   (* //Move Z256 ALM
   "DB_M256M_Scada".tAlm.tS.tS0 := "DB_Z256_Scada".tAlm.tS.tS0;
   "DB_Z256_Scada".tAlm.tS.tS0.x0 := "DB_Z256_Scada".tAlm.tS.tS0.x0;
   "DB_Z256_Scada".tAlm.tS.tS0.x1 := "DB_Z256_Scada".tAlm.tS.tS0.x1;
   "DB_Z256_Scada".tAlm.tS.tS0.x2 := "DB_Z256_Scada".tAlm.tS.tS0.x2;
   "DB_Z256_Scada".tAlm.tS.tS0.x3 := "DB_Z256_Scada".tAlm.tS.tS0.x3;
   "DB_Z256_Scada".tAlm.tS.tS0.x4 := "DB_Z256_Scada".tAlm.tS.tS0.x4;
   "DB_Z256_Scada".tAlm.tS.tS0.x5 := "DB_Z256_Scada".tAlm.tS.tS0.x5;
   "DB_Z256_Scada".tAlm.tS.tS0.x6 := "DB_Z256_Scada".tAlm.tS.tS0.x6;
   "DB_Z256_Scada".tAlm.tS.tS0.x7 := "DB_Z256_Scada".tAlm.tS.tS0.x7;
   "DB_Z256_Scada".tAlm.tS.tS0.x8 := "DB_Z256_Scada".tAlm.tS.tS0.x8;

   "DB_Z256_Scada".tAlm.tS.tS0.x9 := "DB_Z256_Scada".tAlm.tS.tS0.x9;
   "DB_Z256_Scada".tAlm.tS.tS0.x10 := "DB_Z256_Scada".tAlm.tS.tS0.x10;
   "DB_Z256_Scada".tAlm.tS.tS0.x11 := "DB_Z256_Scada".tAlm.tS.tS0.x11;
   "DB_Z256_Scada".tAlm.tS.tS0.x12 := "DB_Z256_Scada".tAlm.tS.tS0.x12;
   "DB_Z256_Scada".tAlm.tS.tS0.x13 := "DB_Z256_Scada".tAlm.tS.tS0.x13;
   "DB_Z256_Scada".tAlm.tS.tS0.x14 := "DB_Z256_Scada".tAlm.tS.tS0.x14;
   "DB_Z256_Scada".tAlm.tS.tS0.x15 := "DB_Z256_Scada".tAlm.tS.tS0.x15;
   "DB_Z256_Scada".tAlm.tS.tS0.x16 := "DB_Z256_Scada".tAlm.tS.tS0.x16;
   "DB_Z256_Scada".tAlm.tS.tS0.x17 := "DB_Z256_Scada".tAlm.tS.tS0.x17;

   "DB_Z256_Scada".tAlm.tS.tS0.x18 := "DB_Z256_Scada".tAlm.tS.tS0.x18;
   "DB_Z256_Scada".tAlm.tS.tS0.x19 := "DB_Z256_Scada".tAlm.tS.tS0.x19;
   "DB_Z256_Scada".tAlm.tS.tS0.x20 := "DB_Z256_Scada".tAlm.tS.tS0.x20;
   "DB_Z256_Scada".tAlm.tS.tS0.x21 := "DB_Z256_Scada".tAlm.tS.tS0.x21;
   "DB_Z256_Scada".tAlm.tS.tS0.x22 := "DB_Z256_Scada".tAlm.tS.tS0.x22;
   "DB_Z256_Scada".tAlm.tS.tS0.x23 := "DB_Z256_Scada".tAlm.tS.tS0.x23;
   "DB_Z256_Scada".tAlm.tS.tS0.x24 := "DB_Z256_Scada".tAlm.tS.tS0.x24;
   "DB_Z256_Scada".tAlm.tS.tS0.x25 := "DB_Z256_Scada".tAlm.tS.tS0.x25;
   "DB_Z256_Scada".tAlm.tS.tS0.x26 := "DB_Z256_Scada".tAlm.tS.tS0.x26;
   "DB_Z256_Scada".tAlm.tS.tS0.x27 := "DB_Z256_Scada".tAlm.tS.tS0.x27;
   "DB_Z256_Scada".tAlm.tS.tS0.x28 := "DB_Z256_Scada".tAlm.tS.tS0.x28;
   "DB_Z256_Scada".tAlm.tS.tS0.x29 := "DB_Z256_Scada".tAlm.tS.tS0.x29;
   "DB_Z256_Scada".tAlm.tS.tS0.x30 := "DB_Z256_Scada".tAlm.tS.tS0.x30;
   "DB_Z256_Scada".tAlm.tS.tS0.x31 := "DB_Z256_Scada".tAlm.tS.tS0.x31; *)


    //Move M256M MOVEMENTS HMR
    //H1
   "DB_M256M_Scada".tHMR.tManCmd.xManJogForwardFdbk_H1 := "M256_Manag_IDB".M256M_IDB[0].tHMR.tManCmd.xMan_JogForwardFdbk;
   "DB_M256M_Scada".tHMR.tManCmd.xManJogBackwardFdbk_H1 := "M256_Manag_IDB".M256M_IDB[0].tHMR.tManCmd.xMan_JogBackwardFdbk;
   "DB_M256M_Scada".tHMR.iCodeAlarm_H1 := "M256_Manag_IDB".M256M_IDB[0].tHMR.iCodeAlarm;
   "DB_M256M_Scada".tHMR.dHeadActualPositions_cmm_H1 := "M256_Manag_IDB".M256M_IDB[0].tHMR.dHeadActualPositions_cmm;
   "DB_M256M_Scada".tHMR.dHeadHomePositions_cmm_H1 := "M256_Manag_IDB".M256M_IDB[0].tHMR.dHeadHomePositions_cmm;
   "DB_M256M_Scada".tHMR.dHeadMoveStatus_H1 := "M256_Manag_IDB".M256M_IDB[0].tHMR.rgdHeadMoveStatus;
   //H2 
   "DB_M256M_Scada".tHMR.tManCmd.xManJogBackwardFdbk_H2 := "M256_Manag_IDB".M256M_IDB[1].tHMR.tManCmd.xMan_JogForwardFdbk;
   "DB_M256M_Scada".tHMR.tManCmd.xManJogBackwardFdbk_H2 := "M256_Manag_IDB".M256M_IDB[1].tHMR.tManCmd.xMan_JogBackwardFdbk;
   "DB_M256M_Scada".tHMR.iCodeAlarm_H2 := "M256_Manag_IDB".M256M_IDB[1].tHMR.iCodeAlarm;
   "DB_M256M_Scada".tHMR.dHeadActualPositions_cmm_H2 := "M256_Manag_IDB".M256M_IDB[1].tHMR.dHeadActualPositions_cmm;
   "DB_M256M_Scada".tHMR.dHeadHomePositions_cmm_H2 := "M256_Manag_IDB".M256M_IDB[1].tHMR.dHeadHomePositions_cmm;
   "DB_M256M_Scada".tHMR.dHeadMoveStatus_H2 := "M256_Manag_IDB".M256M_IDB[1].tHMR.rgdHeadMoveStatus;
   //H3 
   "DB_M256M_Scada".tHMR.tManCmd.xManJogForwardFdbk_H3 :="M256_Manag_IDB".M256M_IDB[2].tHMR.tManCmd.xMan_JogForwardFdbk;
   "DB_M256M_Scada".tHMR.tManCmd.xManJogBackwardFdbk_H3 := "M256_Manag_IDB".M256M_IDB[2].tHMR.tManCmd.xMan_JogBackwardFdbk;
   "DB_M256M_Scada".tHMR.iCodeAlarm_H3 := "M256_Manag_IDB".M256M_IDB[2].tHMR.iCodeAlarm;
   "DB_M256M_Scada".tHMR.dHeadActualPositions_cmm_H3 := "M256_Manag_IDB".M256M_IDB[2].tHMR.dHeadActualPositions_cmm;
   "DB_M256M_Scada".tHMR.dHeadHomePositions_cmm_H3 := "M256_Manag_IDB".M256M_IDB[2].tHMR.dHeadHomePositions_cmm;
   "DB_M256M_Scada".tHMR.dHeadMoveStatus_H3 := "M256_Manag_IDB".M256M_IDB[2].tHMR.rgdHeadMoveStatus;
   //H4 
   "DB_M256M_Scada".tHMR.tManCmd.xManJogForwardFdbk_H4:= "M256_Manag_IDB".M256M_IDB[3].tHMR.tManCmd.xMan_JogForwardFdbk;
   "DB_M256M_Scada".tHMR.tManCmd.xManJogBackwardFdbk_H4 := "M256_Manag_IDB".M256M_IDB[3].tHMR.tManCmd.xMan_JogBackwardFdbk;
   "DB_M256M_Scada".tHMR.iCodeAlarm_H4 := "M256_Manag_IDB".M256M_IDB[3].tHMR.iCodeAlarm;
   "DB_M256M_Scada".tHMR.dHeadActualPositions_cmm_H4 := "M256_Manag_IDB".M256M_IDB[3].tHMR.dHeadActualPositions_cmm;
   "DB_M256M_Scada".tHMR.dHeadHomePositions_cmm_H4 := "M256_Manag_IDB".M256M_IDB[3].tHMR.dHeadHomePositions_cmm;
   "DB_M256M_Scada".tHMR.dHeadMoveStatus_H4 := "M256_Manag_IDB".M256M_IDB[3].tHMR.rgdHeadMoveStatus;
   "DB_M256M_Scada".tHMR.iCodeAlarm_H4 := "M256_Manag_IDB".M256M_IDB[3].tHMR.iCodeAlarm;
   //H5
   "DB_M256M_Scada".tHMR.tManCmd.xManJogForwardFdbk_H5 := "M256_Manag_IDB".M256M_IDB[4].tHMR.tManCmd.xMan_JogForwardFdbk;
   "DB_M256M_Scada".tHMR.tManCmd.xManJogBackwardFdbk_H5:= "M256_Manag_IDB".M256M_IDB[4].tHMR.tManCmd.xMan_JogBackwardFdbk;
   "DB_M256M_Scada".tHMR.iCodeAlarm_H5 := "M256_Manag_IDB".M256M_IDB[4].tHMR.iCodeAlarm;
   "DB_M256M_Scada".tHMR.dHeadActualPositions_cmm_H5 := "M256_Manag_IDB".M256M_IDB[4].tHMR.dHeadActualPositions_cmm;
   "DB_M256M_Scada".tHMR.dHeadHomePositions_cmm_H5 := "M256_Manag_IDB".M256M_IDB[4].tHMR.dHeadHomePositions_cmm;
   "DB_M256M_Scada".tHMR.dHeadMoveStatus_H5 := "M256_Manag_IDB".M256M_IDB[4].tHMR.rgdHeadMoveStatus;
   //H6 
   "DB_M256M_Scada".tHMR.tManCmd.xManJogForwardFdbk_H6 := "M256_Manag_IDB".M256M_IDB[5].tHMR.tManCmd.xMan_JogForwardFdbk;
   "DB_M256M_Scada".tHMR.tManCmd.xManJogBackwardFdbk_H6 := "M256_Manag_IDB".M256M_IDB[5].tHMR.tManCmd.xMan_JogBackwardFdbk;
   "DB_M256M_Scada".tHMR.iCodeAlarm_H6 := "M256_Manag_IDB".M256M_IDB[5].tHMR.iCodeAlarm;
   "DB_M256M_Scada".tHMR.dHeadActualPositions_cmm_H6 := "M256_Manag_IDB".M256M_IDB[5].tHMR.dHeadActualPositions_cmm;
   "DB_M256M_Scada".tHMR.dHeadHomePositions_cmm_H6 := "M256_Manag_IDB".M256M_IDB[5].tHMR.dHeadHomePositions_cmm;
   "DB_M256M_Scada".tHMR.dHeadMoveStatus_H6 := "M256_Manag_IDB".M256M_IDB[5].tHMR.rgdHeadMoveStatus;
   //H7 
   "DB_M256M_Scada".tHMR.tManCmd.xManJogForwardFdbk_H7 := "M256_Manag_IDB".M256M_IDB[6].tHMR.tManCmd.xMan_JogForwardFdbk;
   "DB_M256M_Scada".tHMR.tManCmd.xManJogBackwardFdbk_H7 := "M256_Manag_IDB".M256M_IDB[6].tHMR.tManCmd.xMan_JogBackwardFdbk;
   "DB_M256M_Scada".tHMR.iCodeAlarm_H7 := "M256_Manag_IDB".M256M_IDB[6].tHMR.iCodeAlarm;
   "DB_M256M_Scada".tHMR.dHeadActualPositions_cmm_H7 := "M256_Manag_IDB".M256M_IDB[6].tHMR.dHeadActualPositions_cmm;
   "DB_M256M_Scada".tHMR.dHeadHomePositions_cmm_H7 := "M256_Manag_IDB".M256M_IDB[6].tHMR.dHeadHomePositions_cmm;
   "DB_M256M_Scada".tHMR.dHeadMoveStatus_H7 := "M256_Manag_IDB".M256M_IDB[6].tHMR.rgdHeadMoveStatus;
   //H8 
   "DB_M256M_Scada".tHMR.tManCmd.xManJogForwardFdbk_H8 := "M256_Manag_IDB".M256M_IDB[7].tHMR.tManCmd.xMan_JogForwardFdbk;
   "DB_M256M_Scada".tHMR.tManCmd.xManJogBackwardFdbk_H8 := "M256_Manag_IDB".M256M_IDB[7].tHMR.tManCmd.xMan_JogBackwardFdbk;
   "DB_M256M_Scada".tHMR.iCodeAlarm_H8 := "M256_Manag_IDB".M256M_IDB[7].tHMR.iCodeAlarm;
   "DB_M256M_Scada".tHMR.dHeadActualPositions_cmm_H8 := "M256_Manag_IDB".M256M_IDB[7].tHMR.dHeadActualPositions_cmm;
   "DB_M256M_Scada".tHMR.dHeadHomePositions_cmm_H8 := "M256_Manag_IDB".M256M_IDB[7].tHMR.dHeadHomePositions_cmm;
   "DB_M256M_Scada".tHMR.dHeadMoveStatus_H8 := "M256_Manag_IDB".M256M_IDB[7].tHMR.rgdHeadMoveStatus;


       //Move MOVEMENTS HMW

       //H1
       "M256_Manag_IDB".M256M_IDB[0].tHMW.dHeadHomePositions_cmm := "DB_M256M_Scada".tHMW.dHeadHomePositions_cmm_H1;
       "M256_Manag_IDB".M256M_IDB[0].tHMW.xBrakeEngageHeads := "DB_M256M_Scada".tHMW.xBrakeRealeaseHead_H1;
       "M256_Manag_IDB".M256M_IDB[0].tHMW.xBrakeRealeaseHeads := "DB_M256M_Scada".tHMW.xBrakeEngageHeads_H1;
       "M256_Manag_IDB".M256M_IDB[0].tHMW.xUpdateHomeHead := "DB_M256M_Scada".tHMW.xUpdateHomeHead_H1;
       "M256_Manag_IDB".M256M_IDB[0].tHMW.tManCmd.xMan_JogBackward := "DB_M256M_Scada".tHMW.tManCmd.xMan_JogBackward_H1;
       "M256_Manag_IDB".M256M_IDB[0].tHMW.tManCmd.xMan_JogForward := "DB_M256M_Scada".tHMW.tManCmd.xMan_JogForward_H1;
       //H2
       "M256_Manag_IDB".M256M_IDB[1].tHMW.dHeadHomePositions_cmm := "DB_M256M_Scada".tHMW.dHeadHomePositions_cmm_H2;
       "M256_Manag_IDB".M256M_IDB[1].tHMW.xBrakeEngageHeads := "DB_M256M_Scada".tHMW.xBrakeRealeaseHead_H2;
       "M256_Manag_IDB".M256M_IDB[1].tHMW.xBrakeRealeaseHeads := "DB_M256M_Scada".tHMW.xBrakeEngageHeads_H2;
       "M256_Manag_IDB".M256M_IDB[1].tHMW.xUpdateHomeHead := "DB_M256M_Scada".tHMW.xUpdateHomeHead_H2;
       "M256_Manag_IDB".M256M_IDB[1].tHMW.tManCmd.xMan_JogBackward := "DB_M256M_Scada".tHMW.tManCmd.xMan_JogBackward_H2;
       "M256_Manag_IDB".M256M_IDB[1].tHMW.tManCmd.xMan_JogForward := "DB_M256M_Scada".tHMW.tManCmd.xMan_JogForward_H2;
       //H3
       "M256_Manag_IDB".M256M_IDB[2].tHMW.dHeadHomePositions_cmm := "DB_M256M_Scada".tHMW.dHeadHomePositions_cmm_H3;
       "M256_Manag_IDB".M256M_IDB[2].tHMW.xBrakeEngageHeads := "DB_M256M_Scada".tHMW.xBrakeRealeaseHead_H3;
       "M256_Manag_IDB".M256M_IDB[2].tHMW.xBrakeRealeaseHeads := "DB_M256M_Scada".tHMW.xBrakeEngageHeads_H3;
       "M256_Manag_IDB".M256M_IDB[2].tHMW.xUpdateHomeHead := "DB_M256M_Scada".tHMW.xUpdateHomeHead_H3;
       "M256_Manag_IDB".M256M_IDB[2].tHMW.tManCmd.xMan_JogBackward := "DB_M256M_Scada".tHMW.tManCmd.xMan_JogBackward_H3;
       "M256_Manag_IDB".M256M_IDB[2].tHMW.tManCmd.xMan_JogForward := "DB_M256M_Scada".tHMW.tManCmd.xMan_JogForward_H3;
       //H4
       "M256_Manag_IDB".M256M_IDB[3].tHMW.dHeadHomePositions_cmm := "DB_M256M_Scada".tHMW.dHeadHomePositions_cmm_H4;
       "M256_Manag_IDB".M256M_IDB[3].tHMW.xBrakeEngageHeads := "DB_M256M_Scada".tHMW.xBrakeRealeaseHead_H4;
       "M256_Manag_IDB".M256M_IDB[3].tHMW.xBrakeRealeaseHeads := "DB_M256M_Scada".tHMW.xBrakeEngageHeads_H4;
       "M256_Manag_IDB".M256M_IDB[3].tHMW.xUpdateHomeHead := "DB_M256M_Scada".tHMW.xUpdateHomeHead_H4;
       "M256_Manag_IDB".M256M_IDB[3].tHMW.tManCmd.xMan_JogBackward := "DB_M256M_Scada".tHMW.tManCmd.xMan_JogBackward_H4;
       "M256_Manag_IDB".M256M_IDB[3].tHMW.tManCmd.xMan_JogForward := "DB_M256M_Scada".tHMW.tManCmd.xMan_JogForward_H4;
       //H5
       "M256_Manag_IDB".M256M_IDB[4].tHMW.dHeadHomePositions_cmm := "DB_M256M_Scada".tHMW.dHeadHomePositions_cmm_H5;
       "M256_Manag_IDB".M256M_IDB[4].tHMW.xBrakeEngageHeads := "DB_M256M_Scada".tHMW.xBrakeRealeaseHead_H5;
       "M256_Manag_IDB".M256M_IDB[4].tHMW.xBrakeRealeaseHeads := "DB_M256M_Scada".tHMW.xBrakeEngageHeads_H5;
       "M256_Manag_IDB".M256M_IDB[4].tHMW.xUpdateHomeHead := "DB_M256M_Scada".tHMW.xUpdateHomeHead_H5;
       "M256_Manag_IDB".M256M_IDB[4].tHMW.tManCmd.xMan_JogBackward := "DB_M256M_Scada".tHMW.tManCmd.xMan_JogBackward_H5;
       "M256_Manag_IDB".M256M_IDB[4].tHMW.tManCmd.xMan_JogForward := "DB_M256M_Scada".tHMW.tManCmd.xMan_JogForward_H5;
       //H6
       "M256_Manag_IDB".M256M_IDB[5].tHMW.dHeadHomePositions_cmm := "DB_M256M_Scada".tHMW.dHeadHomePositions_cmm_H6;
       "M256_Manag_IDB".M256M_IDB[5].tHMW.xBrakeEngageHeads := "DB_M256M_Scada".tHMW.xBrakeRealeaseHead_H6;
       "M256_Manag_IDB".M256M_IDB[5].tHMW.xBrakeRealeaseHeads := "DB_M256M_Scada".tHMW.xBrakeEngageHeads_H6;
       "M256_Manag_IDB".M256M_IDB[5].tHMW.xUpdateHomeHead := "DB_M256M_Scada".tHMW.xUpdateHomeHead_H6;
       "M256_Manag_IDB".M256M_IDB[5].tHMW.tManCmd.xMan_JogBackward := "DB_M256M_Scada".tHMW.tManCmd.xMan_JogBackward_H6;
       "M256_Manag_IDB".M256M_IDB[5].tHMW.tManCmd.xMan_JogForward := "DB_M256M_Scada".tHMW.tManCmd.xMan_JogForward_H6;
       //H7
       "M256_Manag_IDB".M256M_IDB[6].tHMW.dHeadHomePositions_cmm := "DB_M256M_Scada".tHMW.dHeadHomePositions_cmm_H7;
       "M256_Manag_IDB".M256M_IDB[6].tHMW.xBrakeEngageHeads := "DB_M256M_Scada".tHMW.xBrakeRealeaseHead_H7;
       "M256_Manag_IDB".M256M_IDB[6].tHMW.xBrakeRealeaseHeads := "DB_M256M_Scada".tHMW.xBrakeEngageHeads_H7;
       "M256_Manag_IDB".M256M_IDB[6].tHMW.xUpdateHomeHead := "DB_M256M_Scada".tHMW.xUpdateHomeHead_H7;
       "M256_Manag_IDB".M256M_IDB[6].tHMW.tManCmd.xMan_JogBackward := "DB_M256M_Scada".tHMW.tManCmd.xMan_JogBackward_H7;
       "M256_Manag_IDB".M256M_IDB[6].tHMW.tManCmd.xMan_JogForward := "DB_M256M_Scada".tHMW.tManCmd.xMan_JogForward_H7;

       //H8
       "M256_Manag_IDB".M256M_IDB[7].tHMW.dHeadHomePositions_cmm := "DB_M256M_Scada".tHMW.dHeadHomePositions_cmm_H8;
       "M256_Manag_IDB".M256M_IDB[7].tHMW.xBrakeEngageHeads := "DB_M256M_Scada".tHMW.xBrakeRealeaseHead_H8;
       "M256_Manag_IDB".M256M_IDB[7].tHMW.xBrakeRealeaseHeads := "DB_M256M_Scada".tHMW.xBrakeEngageHeads_H8;
       "M256_Manag_IDB".M256M_IDB[7].tHMW.xUpdateHomeHead := "DB_M256M_Scada".tHMW.xUpdateHomeHead_H8;
       "M256_Manag_IDB".M256M_IDB[7].tHMW.tManCmd.xMan_JogBackward := "DB_M256M_Scada".tHMW.tManCmd.xMan_JogBackward_H8;
       "M256_Manag_IDB".M256M_IDB[7].tHMW.tManCmd.xMan_JogForward := "DB_M256M_Scada".tHMW.tManCmd.xMan_JogForward_H8;

       //Move MOVEMENTS ALM
       //H1
       "DB_M256M_Scada".tAlm.tS.tS0.x0 := "M256_Manag_IDB".M256M_IDB[0].tALM.tS.x0;
       "DB_M256M_Scada".tAlm.tS.tS0.x1 := "M256_Manag_IDB".M256M_IDB[0].tALM.tS.x1;
       "DB_M256M_Scada".tAlm.tS.tS0.x2 := "M256_Manag_IDB".M256M_IDB[0].tALM.tS.x2;
       "DB_M256M_Scada".tAlm.tS.tS0.x3 := "M256_Manag_IDB".M256M_IDB[0].tALM.tS.x3;
       "DB_M256M_Scada".tAlm.tS.tS0.x4 := "M256_Manag_IDB".M256M_IDB[0].tALM.tS.x4;
       "DB_M256M_Scada".tAlm.tS.tS0.x5 := "M256_Manag_IDB".M256M_IDB[0].tALM.tS.x5;
       "DB_M256M_Scada".tAlm.tS.tS0.x6 := "M256_Manag_IDB".M256M_IDB[0].tALM.tS.x6;
       "DB_M256M_Scada".tAlm.tS.tS0.x7 := "M256_Manag_IDB".M256M_IDB[0].tALM.tS.x7;
       "DB_M256M_Scada".tAlm.tS.tS0.x8 := "M256_Manag_IDB".M256M_IDB[0].tALM.tS.x8;
       //H2
       "DB_M256M_Scada".tAlm.tS.tS0.x9 := "M256_Manag_IDB".M256M_IDB[1].tALM.tS.x0;
       "DB_M256M_Scada".tAlm.tS.tS0.x10 := "M256_Manag_IDB".M256M_IDB[1].tALM.tS.x1;
       "DB_M256M_Scada".tAlm.tS.tS0.x11 := "M256_Manag_IDB".M256M_IDB[1].tALM.tS.x2;
       "DB_M256M_Scada".tAlm.tS.tS0.x12 := "M256_Manag_IDB".M256M_IDB[1].tALM.tS.x3;
       "DB_M256M_Scada".tAlm.tS.tS0.x13 := "M256_Manag_IDB".M256M_IDB[1].tALM.tS.x4;
       "DB_M256M_Scada".tAlm.tS.tS0.x14 := "M256_Manag_IDB".M256M_IDB[1].tALM.tS.x5;
       "DB_M256M_Scada".tAlm.tS.tS0.x15 := "M256_Manag_IDB".M256M_IDB[1].tALM.tS.x6;
       "DB_M256M_Scada".tAlm.tS.tS0.x16 := "M256_Manag_IDB".M256M_IDB[1].tALM.tS.x7;
       "DB_M256M_Scada".tAlm.tS.tS0.x17 := "M256_Manag_IDB".M256M_IDB[1].tALM.tS.x8;
       //H3
       "DB_M256M_Scada".tAlm.tS.tS0.x18 := "M256_Manag_IDB".M256M_IDB[2].tALM.tS.x0;
       "DB_M256M_Scada".tAlm.tS.tS0.x19 := "M256_Manag_IDB".M256M_IDB[2].tALM.tS.x1;
       "DB_M256M_Scada".tAlm.tS.tS0.x20 := "M256_Manag_IDB".M256M_IDB[2].tALM.tS.x2;
       "DB_M256M_Scada".tAlm.tS.tS0.x21 := "M256_Manag_IDB".M256M_IDB[2].tALM.tS.x3;
       "DB_M256M_Scada".tAlm.tS.tS0.x22 := "M256_Manag_IDB".M256M_IDB[2].tALM.tS.x4;
       "DB_M256M_Scada".tAlm.tS.tS0.x23 := "M256_Manag_IDB".M256M_IDB[2].tALM.tS.x5;
       "DB_M256M_Scada".tAlm.tS.tS0.x24 := "M256_Manag_IDB".M256M_IDB[2].tALM.tS.x6;
       "DB_M256M_Scada".tAlm.tS.tS0.x25 := "M256_Manag_IDB".M256M_IDB[2].tALM.tS.x7;
       "DB_M256M_Scada".tAlm.tS.tS0.x26 := "M256_Manag_IDB".M256M_IDB[2].tALM.tS.x8;
       //H4
       "DB_M256M_Scada".tAlm.tS.tS1.x0 := "M256_Manag_IDB".M256M_IDB[3].tALM.tS.x0;
       "DB_M256M_Scada".tAlm.tS.tS1.x1 := "M256_Manag_IDB".M256M_IDB[3].tALM.tS.x1;
       "DB_M256M_Scada".tAlm.tS.tS1.x2 := "M256_Manag_IDB".M256M_IDB[3].tALM.tS.x2;
       "DB_M256M_Scada".tAlm.tS.tS1.x3 := "M256_Manag_IDB".M256M_IDB[3].tALM.tS.x3;
       "DB_M256M_Scada".tAlm.tS.tS1.x4 := "M256_Manag_IDB".M256M_IDB[3].tALM.tS.x4;
       "DB_M256M_Scada".tAlm.tS.tS1.x5 := "M256_Manag_IDB".M256M_IDB[3].tALM.tS.x5;
       "DB_M256M_Scada".tAlm.tS.tS1.x6 := "M256_Manag_IDB".M256M_IDB[3].tALM.tS.x6;
       "DB_M256M_Scada".tAlm.tS.tS1.x7 := "M256_Manag_IDB".M256M_IDB[3].tALM.tS.x7;
       "DB_M256M_Scada".tAlm.tS.tS1.x8 := "M256_Manag_IDB".M256M_IDB[3].tALM.tS.x8;
       //H5
       "DB_M256M_Scada".tAlm.tS.tS1.x9 := "M256_Manag_IDB".M256M_IDB[4].tALM.tS.x0;
       "DB_M256M_Scada".tAlm.tS.tS1.x10 := "M256_Manag_IDB".M256M_IDB[4].tALM.tS.x1;
       "DB_M256M_Scada".tAlm.tS.tS1.x11 := "M256_Manag_IDB".M256M_IDB[4].tALM.tS.x2;
       "DB_M256M_Scada".tAlm.tS.tS1.x12 := "M256_Manag_IDB".M256M_IDB[4].tALM.tS.x3;
       "DB_M256M_Scada".tAlm.tS.tS1.x13 := "M256_Manag_IDB".M256M_IDB[4].tALM.tS.x4;
       "DB_M256M_Scada".tAlm.tS.tS1.x14 := "M256_Manag_IDB".M256M_IDB[4].tALM.tS.x5;
       "DB_M256M_Scada".tAlm.tS.tS1.x15 := "M256_Manag_IDB".M256M_IDB[4].tALM.tS.x6;
       "DB_M256M_Scada".tAlm.tS.tS1.x16 := "M256_Manag_IDB".M256M_IDB[4].tALM.tS.x7;
       "DB_M256M_Scada".tAlm.tS.tS1.x17 := "M256_Manag_IDB".M256M_IDB[4].tALM.tS.x8;
       //H6
       "DB_M256M_Scada".tAlm.tS.tS1.x18 := "M256_Manag_IDB".M256M_IDB[5].tALM.tS.x0;
       "DB_M256M_Scada".tAlm.tS.tS1.x19 := "M256_Manag_IDB".M256M_IDB[5].tALM.tS.x1;
       "DB_M256M_Scada".tAlm.tS.tS1.x20 := "M256_Manag_IDB".M256M_IDB[5].tALM.tS.x2;
       "DB_M256M_Scada".tAlm.tS.tS1.x21 := "M256_Manag_IDB".M256M_IDB[5].tALM.tS.x3;
       "DB_M256M_Scada".tAlm.tS.tS1.x22 := "M256_Manag_IDB".M256M_IDB[5].tALM.tS.x4;
       "DB_M256M_Scada".tAlm.tS.tS1.x23 := "M256_Manag_IDB".M256M_IDB[5].tALM.tS.x5;
       "DB_M256M_Scada".tAlm.tS.tS1.x24 := "M256_Manag_IDB".M256M_IDB[5].tALM.tS.x6;
       "DB_M256M_Scada".tAlm.tS.tS1.x25 := "M256_Manag_IDB".M256M_IDB[5].tALM.tS.x7;
       "DB_M256M_Scada".tAlm.tS.tS1.x26 := "M256_Manag_IDB".M256M_IDB[5].tALM.tS.x8;
       //H7
       "DB_M256M_Scada".tAlm.tS.tS2.x0 := "M256_Manag_IDB".M256M_IDB[6].tALM.tS.x0;
       "DB_M256M_Scada".tAlm.tS.tS2.x1 := "M256_Manag_IDB".M256M_IDB[6].tALM.tS.x1;
       "DB_M256M_Scada".tAlm.tS.tS2.x2 := "M256_Manag_IDB".M256M_IDB[6].tALM.tS.x2;
       "DB_M256M_Scada".tAlm.tS.tS2.x3 := "M256_Manag_IDB".M256M_IDB[6].tALM.tS.x3;
       "DB_M256M_Scada".tAlm.tS.tS2.x4 := "M256_Manag_IDB".M256M_IDB[6].tALM.tS.x4;
       "DB_M256M_Scada".tAlm.tS.tS2.x5 := "M256_Manag_IDB".M256M_IDB[6].tALM.tS.x5;
       "DB_M256M_Scada".tAlm.tS.tS2.x6 := "M256_Manag_IDB".M256M_IDB[6].tALM.tS.x6;
       "DB_M256M_Scada".tAlm.tS.tS2.x7 := "M256_Manag_IDB".M256M_IDB[6].tALM.tS.x7;
       "DB_M256M_Scada".tAlm.tS.tS2.x8 := "M256_Manag_IDB".M256M_IDB[6].tALM.tS.x8;
       //H8
       "DB_M256M_Scada".tAlm.tS.tS2.x9 := "M256_Manag_IDB".M256M_IDB[7].tALM.tS.x0;
       "DB_M256M_Scada".tAlm.tS.tS2.x10 := "M256_Manag_IDB".M256M_IDB[7].tALM.tS.x1;
       "DB_M256M_Scada".tAlm.tS.tS2.x11 := "M256_Manag_IDB".M256M_IDB[7].tALM.tS.x2;
       "DB_M256M_Scada".tAlm.tS.tS2.x12:= "M256_Manag_IDB".M256M_IDB[7].tALM.tS.x3;
       "DB_M256M_Scada".tAlm.tS.tS2.x13 := "M256_Manag_IDB".M256M_IDB[7].tALM.tS.x4;
       "DB_M256M_Scada".tAlm.tS.tS2.x14 := "M256_Manag_IDB".M256M_IDB[7].tALM.tS.x5;
       "DB_M256M_Scada".tAlm.tS.tS2.x15 := "M256_Manag_IDB".M256M_IDB[7].tALM.tS.x6;
       "DB_M256M_Scada".tAlm.tS.tS2.x16 := "M256_Manag_IDB".M256M_IDB[7].tALM.tS.x7;
       "DB_M256M_Scada".tAlm.tS.tS2.x17 := "M256_Manag_IDB".M256M_IDB[7].tALM.tS.x8;


       //Move FIRE HMR
       //H1
       "DB_M256F_Scada".tHMR.dHeadStatus_H1 := "M256_Manag_IDB".M256F_IDB[0].tHMR.dHeadStatus;
       "DB_M256F_Scada".tHMR.rHeadUsage_km_H1 := "M256_Manag_IDB".M256F_IDB[0].tHMR.rHeadUsage_km;
       "DB_M256F_Scada".tHMR.tManCmd.xMan_FireON_Fdbk_H1 := "M256_Manag_IDB".M256F_IDB[0].tHMR.tManCmd.xMan_FireON_Fdbk;
       "DB_M256F_Scada".tHMR.tManCmd.xMan_FireOFF_Fdbk_H1 := "M256_Manag_IDB".M256F_IDB[0].tHMR.tManCmd.xMan_FireOFF_Fdbk;
       "DB_M256F_Scada".tHMR.tManCmd.xMan_OilON_Fdbk_H1 := "M256_Manag_IDB".M256F_IDB[0].tHMR.tManCmd.xMan_OilON_Fdbk;

       //H2
       "DB_M256F_Scada".tHMR.dHeadStatus_H2 := "M256_Manag_IDB".M256F_IDB[1].tHMR.dHeadStatus;
       "DB_M256F_Scada".tHMR.rHeadUsage_km_H2 := "M256_Manag_IDB".M256F_IDB[1].tHMR.rHeadUsage_km;
       "DB_M256F_Scada".tHMR.tManCmd.xMan_FireON_Fdbk_H2 := "M256_Manag_IDB".M256F_IDB[1].tHMR.tManCmd.xMan_FireON_Fdbk;
       "DB_M256F_Scada".tHMR.tManCmd.xMan_FireOFF_Fdbk_H2 := "M256_Manag_IDB".M256F_IDB[1].tHMR.tManCmd.xMan_FireOFF_Fdbk;
       "DB_M256F_Scada".tHMR.tManCmd.xMan_OilON_Fdbk_H2 := "M256_Manag_IDB".M256F_IDB[1].tHMR.tManCmd.xMan_OilON_Fdbk;

       //H3
       "DB_M256F_Scada".tHMR.dHeadStatus_H3 := "M256_Manag_IDB".M256F_IDB[2].tHMR.dHeadStatus;
       "DB_M256F_Scada".tHMR.rHeadUsage_km_H3 := "M256_Manag_IDB".M256F_IDB[2].tHMR.rHeadUsage_km;
       "DB_M256F_Scada".tHMR.tManCmd.xMan_FireON_Fdbk_H3 := "M256_Manag_IDB".M256F_IDB[2].tHMR.tManCmd.xMan_FireON_Fdbk;
       "DB_M256F_Scada".tHMR.tManCmd.xMan_FireOFF_Fdbk_H3 := "M256_Manag_IDB".M256F_IDB[2].tHMR.tManCmd.xMan_FireOFF_Fdbk;
       "DB_M256F_Scada".tHMR.tManCmd.xMan_OilON_Fdbk_H3 := "M256_Manag_IDB".M256F_IDB[2].tHMR.tManCmd.xMan_OilON_Fdbk;
       //H4
       "DB_M256F_Scada".tHMR.dHeadStatus_H4 := "M256_Manag_IDB".M256F_IDB[3].tHMR.dHeadStatus;
       "DB_M256F_Scada".tHMR.rHeadUsage_km_H4 := "M256_Manag_IDB".M256F_IDB[3].tHMR.rHeadUsage_km;
       "DB_M256F_Scada".tHMR.tManCmd.xMan_FireON_Fdbk_H4 := "M256_Manag_IDB".M256F_IDB[3].tHMR.tManCmd.xMan_FireON_Fdbk;
       "DB_M256F_Scada".tHMR.tManCmd.xMan_FireOFF_Fdbk_H4 := "M256_Manag_IDB".M256F_IDB[3].tHMR.tManCmd.xMan_FireOFF_Fdbk;
       "DB_M256F_Scada".tHMR.tManCmd.xMan_OilON_Fdbk_H4 := "M256_Manag_IDB".M256F_IDB[3].tHMR.tManCmd.xMan_OilON_Fdbk;
       //H5
       "DB_M256F_Scada".tHMR.dHeadStatus_H5 := "M256_Manag_IDB".M256F_IDB[4].tHMR.dHeadStatus;
       "DB_M256F_Scada".tHMR.rHeadUsage_km_H5 := "M256_Manag_IDB".M256F_IDB[4].tHMR.rHeadUsage_km;
       "DB_M256F_Scada".tHMR.tManCmd.xMan_FireON_Fdbk_H5 := "M256_Manag_IDB".M256F_IDB[4].tHMR.tManCmd.xMan_FireON_Fdbk;
       "DB_M256F_Scada".tHMR.tManCmd.xMan_FireOFF_Fdbk_H5 := "M256_Manag_IDB".M256F_IDB[4].tHMR.tManCmd.xMan_FireOFF_Fdbk;
       "DB_M256F_Scada".tHMR.tManCmd.xMan_OilON_Fdbk_H5 := "M256_Manag_IDB".M256F_IDB[4].tHMR.tManCmd.xMan_OilON_Fdbk;
       //H6
       "DB_M256F_Scada".tHMR.dHeadStatus_H6 := "M256_Manag_IDB".M256F_IDB[5].tHMR.dHeadStatus;
       "DB_M256F_Scada".tHMR.rHeadUsage_km_H6 := "M256_Manag_IDB".M256F_IDB[5].tHMR.rHeadUsage_km;
       "DB_M256F_Scada".tHMR.tManCmd.xMan_FireON_Fdbk_H6 := "M256_Manag_IDB".M256F_IDB[5].tHMR.tManCmd.xMan_FireON_Fdbk;
       "DB_M256F_Scada".tHMR.tManCmd.xMan_FireOFF_Fdbk_H6 := "M256_Manag_IDB".M256F_IDB[5].tHMR.tManCmd.xMan_FireOFF_Fdbk;
       "DB_M256F_Scada".tHMR.tManCmd.xMan_OilON_Fdbk_H6 := "M256_Manag_IDB".M256F_IDB[5].tHMR.tManCmd.xMan_OilON_Fdbk;
       //H7
       "DB_M256F_Scada".tHMR.dHeadStatus_H7 := "M256_Manag_IDB".M256F_IDB[6].tHMR.dHeadStatus;
       "DB_M256F_Scada".tHMR.rHeadUsage_km_H7 := "M256_Manag_IDB".M256F_IDB[6].tHMR.rHeadUsage_km;
       "DB_M256F_Scada".tHMR.tManCmd.xMan_FireON_Fdbk_H7 := "M256_Manag_IDB".M256F_IDB[6].tHMR.tManCmd.xMan_FireON_Fdbk;
       "DB_M256F_Scada".tHMR.tManCmd.xMan_FireOFF_Fdbk_H7 := "M256_Manag_IDB".M256F_IDB[6].tHMR.tManCmd.xMan_FireOFF_Fdbk;
       "DB_M256F_Scada".tHMR.tManCmd.xMan_OilON_Fdbk_H7 := "M256_Manag_IDB".M256F_IDB[6].tHMR.tManCmd.xMan_OilON_Fdbk;
       //H8
       "DB_M256F_Scada".tHMR.dHeadStatus_H8 := "M256_Manag_IDB".M256F_IDB[7].tHMR.dHeadStatus;
       "DB_M256F_Scada".tHMR.rHeadUsage_km_H8 := "M256_Manag_IDB".M256F_IDB[7].tHMR.rHeadUsage_km;
       "DB_M256F_Scada".tHMR.tManCmd.xMan_FireON_Fdbk_H8 := "M256_Manag_IDB".M256F_IDB[7].tHMR.tManCmd.xMan_FireON_Fdbk;
       "DB_M256F_Scada".tHMR.tManCmd.xMan_FireOFF_Fdbk_H8 := "M256_Manag_IDB".M256F_IDB[7].tHMR.tManCmd.xMan_FireOFF_Fdbk;
       "DB_M256F_Scada".tHMR.tManCmd.xMan_OilON_Fdbk_H8 := "M256_Manag_IDB".M256F_IDB[7].tHMR.tManCmd.xMan_OilON_Fdbk;




       //Move FIRE HMW
       //H1
       "M256_Manag_IDB".M256F_IDB[0].tHMW.dHeadFireONReaction_ms := "DB_M256F_Scada".tHMW.dHeadFireONReaction_ms_H1;
       "M256_Manag_IDB".M256F_IDB[0].tHMW.dHeadFireOFFReaction_ms := "DB_M256F_Scada".tHMW.dHeadFireOFFReaction_ms_H1;
       "M256_Manag_IDB".M256F_IDB[0].tHMW.dHeadOilONDelay_ms := "DB_M256F_Scada".tHMW.dHeadOilONDelay_ms_H1;
       "M256_Manag_IDB".M256F_IDB[0].tHMW.dHeadOilOFFDelay_ms := "DB_M256F_Scada".tHMW.dHeadOilOFFDelay_ms_H1;
       "M256_Manag_IDB".M256F_IDB[0].tHMW.dHeadFireONDelay_cmm := "DB_M256F_Scada".tHMW.dHeadFireONDelay_cmm_H1;
       "M256_Manag_IDB".M256F_IDB[0].tHMW.dHeadFireOFFDelay_cmm := "DB_M256F_Scada".tHMW.dHeadFireOFFDelay_cmm_H1;
       "M256_Manag_IDB".M256F_IDB[0].tHMW.dHeadPressure_mN := "DB_M256F_Scada".tHMW.dHeadPressure_mN_H1;
       "M256_Manag_IDB".M256F_IDB[0].tHMW.xResetUsageCounter := "DB_M256F_Scada".tHMW.xResetUsageCounter_H1;
       "M256_Manag_IDB".M256F_IDB[0].tHMW.tManCmd.xMan_FireON := "DB_M256F_Scada".tHMW.tManCmd.xMan_FireON_H1;
       "M256_Manag_IDB".M256F_IDB[0].tHMW.tManCmd.xMan_FireOFF := "DB_M256F_Scada".tHMW.tManCmd.xMan_FireOFF_H1;
       "M256_Manag_IDB".M256F_IDB[0].tHMW.tManCmd.xMan_OilON := "DB_M256F_Scada".tHMW.tManCmd.xMan_OilON_H1;
       //H2
       "M256_Manag_IDB".M256F_IDB[1].tHMW.dHeadFireONReaction_ms := "DB_M256F_Scada".tHMW.dHeadFireONReaction_ms_H2;
       "M256_Manag_IDB".M256F_IDB[1].tHMW.dHeadFireOFFReaction_ms := "DB_M256F_Scada".tHMW.dHeadFireOFFReaction_ms_H2;
       "M256_Manag_IDB".M256F_IDB[1].tHMW.dHeadOilONDelay_ms := "DB_M256F_Scada".tHMW.dHeadOilONDelay_ms_H2;
       "M256_Manag_IDB".M256F_IDB[1].tHMW.dHeadOilOFFDelay_ms := "DB_M256F_Scada".tHMW.dHeadOilOFFDelay_ms_H2;
       "M256_Manag_IDB".M256F_IDB[1].tHMW.dHeadFireONDelay_cmm := "DB_M256F_Scada".tHMW.dHeadFireONDelay_cmm_H2;
       "M256_Manag_IDB".M256F_IDB[1].tHMW.dHeadFireOFFDelay_cmm := "DB_M256F_Scada".tHMW.dHeadFireOFFDelay_cmm_H2;
       "M256_Manag_IDB".M256F_IDB[1].tHMW.dHeadPressure_mN := "DB_M256F_Scada".tHMW.dHeadPressure_mN_H2;
       "M256_Manag_IDB".M256F_IDB[1].tHMW.xResetUsageCounter := "DB_M256F_Scada".tHMW.xResetUsageCounter_H2;
       "M256_Manag_IDB".M256F_IDB[1].tHMW.tManCmd.xMan_FireON := "DB_M256F_Scada".tHMW.tManCmd.xMan_FireON_H2;
       "M256_Manag_IDB".M256F_IDB[1].tHMW.tManCmd.xMan_FireOFF := "DB_M256F_Scada".tHMW.tManCmd.xMan_FireOFF_H2;
       "M256_Manag_IDB".M256F_IDB[1].tHMW.tManCmd.xMan_OilON := "DB_M256F_Scada".tHMW.tManCmd.xMan_OilON_H2;
       //H3
       "M256_Manag_IDB".M256F_IDB[2].tHMW.dHeadFireONReaction_ms := "DB_M256F_Scada".tHMW.dHeadFireONReaction_ms_H3;
       "M256_Manag_IDB".M256F_IDB[2].tHMW.dHeadFireOFFReaction_ms := "DB_M256F_Scada".tHMW.dHeadFireOFFReaction_ms_H3;
       "M256_Manag_IDB".M256F_IDB[2].tHMW.dHeadOilONDelay_ms := "DB_M256F_Scada".tHMW.dHeadOilONDelay_ms_H3;
       "M256_Manag_IDB".M256F_IDB[2].tHMW.dHeadOilOFFDelay_ms := "DB_M256F_Scada".tHMW.dHeadOilOFFDelay_ms_H3;
       "M256_Manag_IDB".M256F_IDB[2].tHMW.dHeadFireONDelay_cmm := "DB_M256F_Scada".tHMW.dHeadFireONDelay_cmm_H3;
       "M256_Manag_IDB".M256F_IDB[2].tHMW.dHeadFireOFFDelay_cmm := "DB_M256F_Scada".tHMW.dHeadFireOFFDelay_cmm_H3;
       "M256_Manag_IDB".M256F_IDB[2].tHMW.dHeadPressure_mN := "DB_M256F_Scada".tHMW.dHeadPressure_mN_H3;
       "M256_Manag_IDB".M256F_IDB[2].tHMW.xResetUsageCounter := "DB_M256F_Scada".tHMW.xResetUsageCounter_H3;
       "M256_Manag_IDB".M256F_IDB[2].tHMW.tManCmd.xMan_FireON := "DB_M256F_Scada".tHMW.tManCmd.xMan_FireON_H3;
       "M256_Manag_IDB".M256F_IDB[2].tHMW.tManCmd.xMan_FireOFF := "DB_M256F_Scada".tHMW.tManCmd.xMan_FireOFF_H3;
       "M256_Manag_IDB".M256F_IDB[2].tHMW.tManCmd.xMan_OilON := "DB_M256F_Scada".tHMW.tManCmd.xMan_OilON_H3;
       //H4
       "M256_Manag_IDB".M256F_IDB[3].tHMW.dHeadFireONReaction_ms := "DB_M256F_Scada".tHMW.dHeadFireONReaction_ms_H4;
       "M256_Manag_IDB".M256F_IDB[3].tHMW.dHeadFireOFFReaction_ms := "DB_M256F_Scada".tHMW.dHeadFireOFFReaction_ms_H4;
       "M256_Manag_IDB".M256F_IDB[3].tHMW.dHeadOilONDelay_ms := "DB_M256F_Scada".tHMW.dHeadOilONDelay_ms_H4;
       "M256_Manag_IDB".M256F_IDB[3].tHMW.dHeadOilOFFDelay_ms := "DB_M256F_Scada".tHMW.dHeadOilOFFDelay_ms_H4;
       "M256_Manag_IDB".M256F_IDB[3].tHMW.dHeadFireONDelay_cmm := "DB_M256F_Scada".tHMW.dHeadFireONDelay_cmm_H4;
       "M256_Manag_IDB".M256F_IDB[3].tHMW.dHeadFireOFFDelay_cmm := "DB_M256F_Scada".tHMW.dHeadFireOFFDelay_cmm_H4;
       "M256_Manag_IDB".M256F_IDB[3].tHMW.dHeadPressure_mN := "DB_M256F_Scada".tHMW.dHeadPressure_mN_H4;
       "M256_Manag_IDB".M256F_IDB[3].tHMW.xResetUsageCounter := "DB_M256F_Scada".tHMW.xResetUsageCounter_H4;
       "M256_Manag_IDB".M256F_IDB[3].tHMW.tManCmd.xMan_FireON := "DB_M256F_Scada".tHMW.tManCmd.xMan_FireON_H4;
       "M256_Manag_IDB".M256F_IDB[3].tHMW.tManCmd.xMan_FireOFF := "DB_M256F_Scada".tHMW.tManCmd.xMan_FireOFF_H4;
       "M256_Manag_IDB".M256F_IDB[3].tHMW.tManCmd.xMan_OilON := "DB_M256F_Scada".tHMW.tManCmd.xMan_OilON_H4;
       //H5
       "M256_Manag_IDB".M256F_IDB[4].tHMW.dHeadFireONReaction_ms := "DB_M256F_Scada".tHMW.dHeadFireONReaction_ms_H5;
       "M256_Manag_IDB".M256F_IDB[4].tHMW.dHeadFireOFFReaction_ms := "DB_M256F_Scada".tHMW.dHeadFireOFFReaction_ms_H5;
       "M256_Manag_IDB".M256F_IDB[4].tHMW.dHeadOilONDelay_ms := "DB_M256F_Scada".tHMW.dHeadOilONDelay_ms_H5;
       "M256_Manag_IDB".M256F_IDB[4].tHMW.dHeadOilOFFDelay_ms := "DB_M256F_Scada".tHMW.dHeadOilOFFDelay_ms_H5;
       "M256_Manag_IDB".M256F_IDB[4].tHMW.dHeadFireONDelay_cmm := "DB_M256F_Scada".tHMW.dHeadFireONDelay_cmm_H5;
       "M256_Manag_IDB".M256F_IDB[4].tHMW.dHeadFireOFFDelay_cmm := "DB_M256F_Scada".tHMW.dHeadFireOFFDelay_cmm_H5;
       "M256_Manag_IDB".M256F_IDB[4].tHMW.dHeadPressure_mN := "DB_M256F_Scada".tHMW.dHeadPressure_mN_H5;
       "M256_Manag_IDB".M256F_IDB[4].tHMW.xResetUsageCounter := "DB_M256F_Scada".tHMW.xResetUsageCounter_H5;
       "M256_Manag_IDB".M256F_IDB[4].tHMW.tManCmd.xMan_FireON := "DB_M256F_Scada".tHMW.tManCmd.xMan_FireON_H5;
       "M256_Manag_IDB".M256F_IDB[4].tHMW.tManCmd.xMan_FireOFF := "DB_M256F_Scada".tHMW.tManCmd.xMan_FireOFF_H5;
       "M256_Manag_IDB".M256F_IDB[4].tHMW.tManCmd.xMan_OilON := "DB_M256F_Scada".tHMW.tManCmd.xMan_OilON_H5;
       //H6
       "M256_Manag_IDB".M256F_IDB[5].tHMW.dHeadFireONReaction_ms := "DB_M256F_Scada".tHMW.dHeadFireONReaction_ms_H6;
       "M256_Manag_IDB".M256F_IDB[5].tHMW.dHeadFireOFFReaction_ms := "DB_M256F_Scada".tHMW.dHeadFireOFFReaction_ms_H6;
       "M256_Manag_IDB".M256F_IDB[5].tHMW.dHeadOilONDelay_ms := "DB_M256F_Scada".tHMW.dHeadOilONDelay_ms_H6;
       "M256_Manag_IDB".M256F_IDB[5].tHMW.dHeadOilOFFDelay_ms := "DB_M256F_Scada".tHMW.dHeadOilOFFDelay_ms_H6;
       "M256_Manag_IDB".M256F_IDB[5].tHMW.dHeadFireONDelay_cmm := "DB_M256F_Scada".tHMW.dHeadFireONDelay_cmm_H6;
       "M256_Manag_IDB".M256F_IDB[5].tHMW.dHeadFireOFFDelay_cmm := "DB_M256F_Scada".tHMW.dHeadFireOFFDelay_cmm_H6;
       "M256_Manag_IDB".M256F_IDB[5].tHMW.dHeadPressure_mN := "DB_M256F_Scada".tHMW.dHeadPressure_mN_H6;
       "M256_Manag_IDB".M256F_IDB[5].tHMW.xResetUsageCounter := "DB_M256F_Scada".tHMW.xResetUsageCounter_H6;
       "M256_Manag_IDB".M256F_IDB[5].tHMW.tManCmd.xMan_FireON := "DB_M256F_Scada".tHMW.tManCmd.xMan_FireON_H6;
       "M256_Manag_IDB".M256F_IDB[5].tHMW.tManCmd.xMan_FireOFF := "DB_M256F_Scada".tHMW.tManCmd.xMan_FireOFF_H6;
       "M256_Manag_IDB".M256F_IDB[5].tHMW.tManCmd.xMan_OilON := "DB_M256F_Scada".tHMW.tManCmd.xMan_OilON_H6;
       //H7
       "M256_Manag_IDB".M256F_IDB[6].tHMW.dHeadFireONReaction_ms := "DB_M256F_Scada".tHMW.dHeadFireONReaction_ms_H7;
       "M256_Manag_IDB".M256F_IDB[6].tHMW.dHeadFireOFFReaction_ms := "DB_M256F_Scada".tHMW.dHeadFireOFFReaction_ms_H7;
       "M256_Manag_IDB".M256F_IDB[6].tHMW.dHeadOilONDelay_ms := "DB_M256F_Scada".tHMW.dHeadOilONDelay_ms_H7;
       "M256_Manag_IDB".M256F_IDB[6].tHMW.dHeadOilOFFDelay_ms := "DB_M256F_Scada".tHMW.dHeadOilOFFDelay_ms_H7;
       "M256_Manag_IDB".M256F_IDB[6].tHMW.dHeadFireONDelay_cmm := "DB_M256F_Scada".tHMW.dHeadFireONDelay_cmm_H7;
       "M256_Manag_IDB".M256F_IDB[6].tHMW.dHeadFireOFFDelay_cmm := "DB_M256F_Scada".tHMW.dHeadFireOFFDelay_cmm_H7;
       "M256_Manag_IDB".M256F_IDB[6].tHMW.dHeadPressure_mN := "DB_M256F_Scada".tHMW.dHeadPressure_mN_H7;
       "M256_Manag_IDB".M256F_IDB[6].tHMW.xResetUsageCounter := "DB_M256F_Scada".tHMW.xResetUsageCounter_H7;
       "M256_Manag_IDB".M256F_IDB[6].tHMW.tManCmd.xMan_FireON := "DB_M256F_Scada".tHMW.tManCmd.xMan_FireON_H7;
       "M256_Manag_IDB".M256F_IDB[6].tHMW.tManCmd.xMan_FireOFF := "DB_M256F_Scada".tHMW.tManCmd.xMan_FireOFF_H7;
       "M256_Manag_IDB".M256F_IDB[6].tHMW.tManCmd.xMan_OilON := "DB_M256F_Scada".tHMW.tManCmd.xMan_OilON_H7;
       //H8
       "M256_Manag_IDB".M256F_IDB[7].tHMW.dHeadFireONReaction_ms := "DB_M256F_Scada".tHMW.dHeadFireONReaction_ms_H8;
       "M256_Manag_IDB".M256F_IDB[7].tHMW.dHeadFireOFFReaction_ms := "DB_M256F_Scada".tHMW.dHeadFireOFFReaction_ms_H8;
       "M256_Manag_IDB".M256F_IDB[7].tHMW.dHeadOilONDelay_ms := "DB_M256F_Scada".tHMW.dHeadOilONDelay_ms_H8;
       "M256_Manag_IDB".M256F_IDB[7].tHMW.dHeadOilOFFDelay_ms := "DB_M256F_Scada".tHMW.dHeadOilOFFDelay_ms_H8;
       "M256_Manag_IDB".M256F_IDB[7].tHMW.dHeadFireONDelay_cmm := "DB_M256F_Scada".tHMW.dHeadFireONDelay_cmm_H8;
       "M256_Manag_IDB".M256F_IDB[7].tHMW.dHeadFireOFFDelay_cmm := "DB_M256F_Scada".tHMW.dHeadFireOFFDelay_cmm_H8;
       "M256_Manag_IDB".M256F_IDB[7].tHMW.dHeadPressure_mN := "DB_M256F_Scada".tHMW.dHeadPressure_mN_H8;
       "M256_Manag_IDB".M256F_IDB[7].tHMW.xResetUsageCounter := "DB_M256F_Scada".tHMW.xResetUsageCounter_H8;
       "M256_Manag_IDB".M256F_IDB[7].tHMW.tManCmd.xMan_FireON := "DB_M256F_Scada".tHMW.tManCmd.xMan_FireON_H8;
       "M256_Manag_IDB".M256F_IDB[7].tHMW.tManCmd.xMan_FireOFF := "DB_M256F_Scada".tHMW.tManCmd.xMan_FireOFF_H8;
       "M256_Manag_IDB".M256F_IDB[7].tHMW.tManCmd.xMan_OilON := "DB_M256F_Scada".tHMW.tManCmd.xMan_OilON_H8;

       //Move FIRE ALM
       "DB_M256F_Scada".tAlm.tF:="M256_Manag_IDB".M256F_IDB[0].tALM.tF;

       "DB_M256F_Scada".tAlm.tW := "M256_Manag_IDB".M256F_IDB[0].tALM.tW;